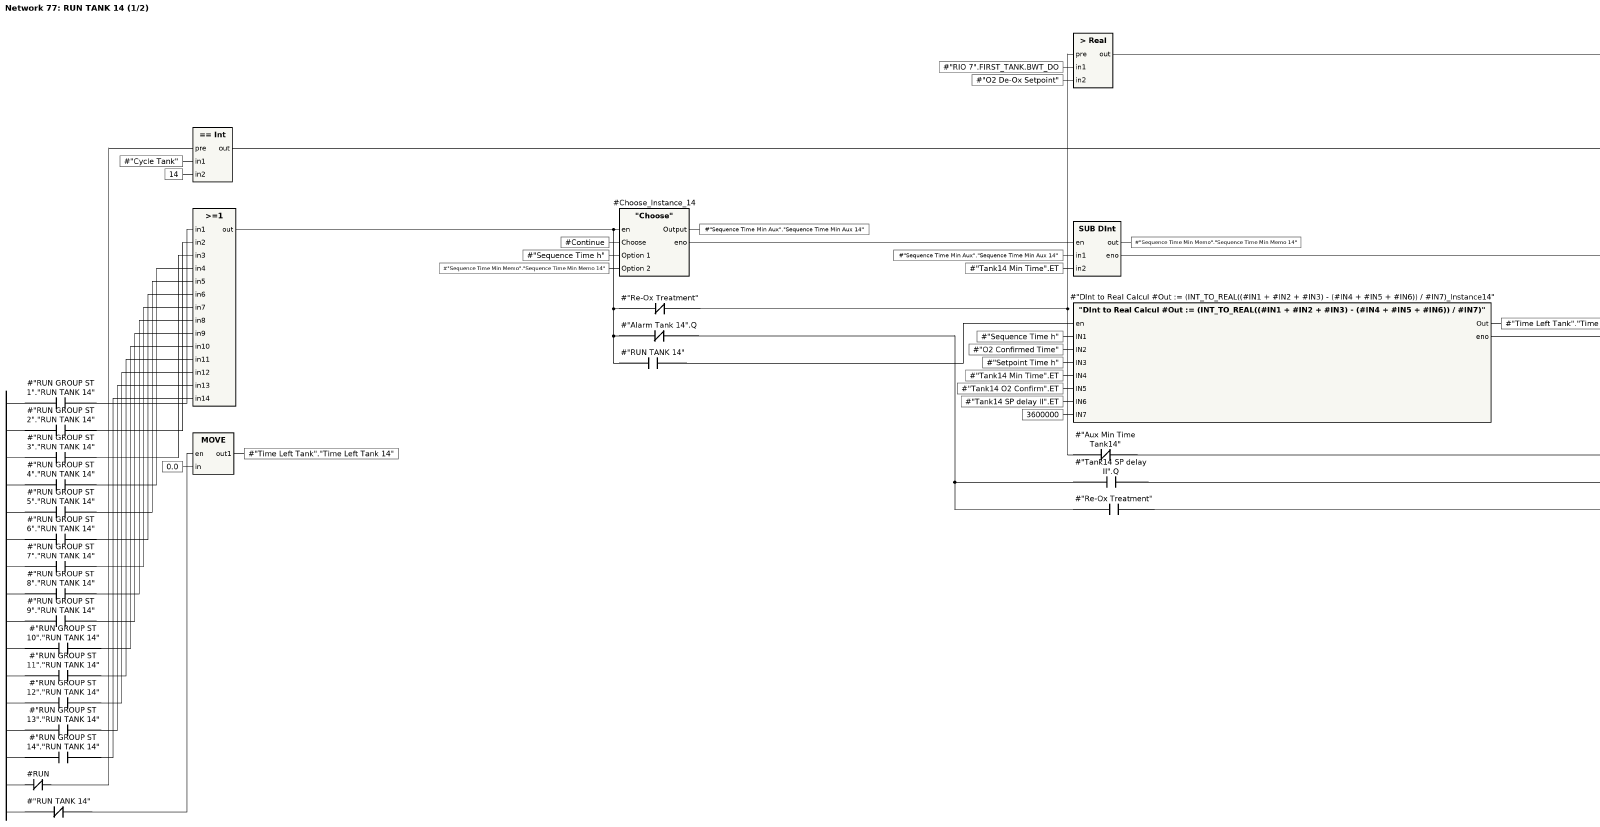
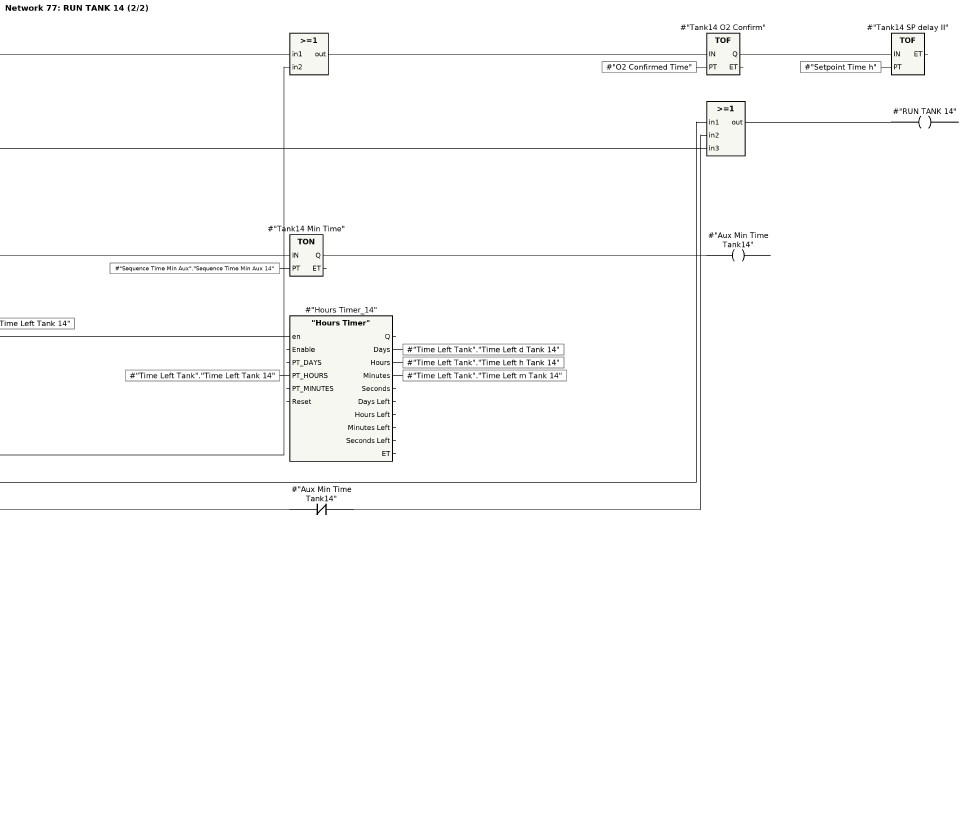
   #_w1 := #"RUN GROUP ST 1"."RUN TANK 14" OR #"RUN GROUP ST 2"."RUN TANK 14" OR #"RUN GROUP ST 3"."RUN TANK 14" OR #"RUN GROUP ST 4"."RUN TANK 14" OR #"RUN GROUP ST 5"."RUN TANK 14" OR #"RUN GROUP ST 6"."RUN TANK 14" OR #"RUN GROUP ST 7"."RUN TANK 14" OR #"RUN GROUP ST 8"."RUN TANK 14" OR #"RUN GROUP ST 9"."RUN TANK 14" OR #"RUN GROUP ST 10"."RUN TANK 14" OR #"RUN GROUP ST 11"."RUN TANK 14" OR #"RUN GROUP ST 12"."RUN TANK 14" OR #"RUN GROUP ST 13"."RUN TANK 14" OR #"RUN GROUP ST 14"."RUN TANK 14";
   #Choose_Instance_14(EN := #_w1,   // "Choose"
                       Choose := #Continue,
                       "Option 1" := #"Sequence Time h",
                       "Option 2" := #"Sequence Time Min Memo"."Sequence Time Min Memo 14",
                       Output => #"Sequence Time Min Aux"."Sequence Time Min Aux 14",
                       ENO => #_w2);
   IF #_w2 THEN
       #"Sequence Time Min Memo"."Sequence Time Min Memo 14" := #"Sequence Time Min Aux"."Sequence Time Min Aux 14" - #"Tank14 Min Time".ET;   // Memory of remained time for use to continue
   END_IF;
   #"Tank14 Min Time"(IN := #_w2, PT := #"Sequence Time Min Aux"."Sequence Time Min Aux 14");   // TON
   #"Aux Min Time Tank14" := #"Tank14 Min Time".Q;
   #"Tank14 O2 Confirm"(IN := #_w1 AND NOT #"Re-Ox Treatment" AND ((#"RIO 7".FIRST_TANK.BWT_DO > #"O2 De-Ox Setpoint") OR NOT #"Aux Min Time Tank14"),   // TOF
                        PT := #"O2 Confirmed Time");
   #"Tank14 SP delay II"(IN := #"Tank14 O2 Confirm".Q, PT := #"Setpoint Time h");   // TOF
   #"DInt to Real Calcul #Out := (INT_TO_REAL((#IN1 + #IN2 + #IN3) - (#IN4 + #IN5 + #IN6)) / #IN7)_Instance14"(EN := #_w1 AND #"RUN TANK 14",   // "DInt to Real Calcul #Out := (INT_TO_REAL((#IN1 + #IN2 + #IN3) - (#IN4 + #IN5 + #IN6)) / #IN7)"
                           IN1 := #"Sequence Time h",
                           IN2 := #"O2 Confirmed Time",
                           IN3 := #"Setpoint Time h",
                           IN4 := #"Tank14 Min Time".ET,
                           IN5 := #"Tank14 O2 Confirm".ET,
                           IN6 := #"Tank14 SP delay II".ET,
                           IN7 := 3600000,
                           Out => #"Time Left Tank"."Time Left Tank 14",
                           ENO => #_w3);
   IF #_w3 THEN
       #"Hours Timer_14"(PT_HOURS := #"Time Left Tank"."Time Left Tank 14",   // "Hours Timer"
                         Days => #"Time Left Tank"."Time Left d Tank 14",
                         Hours => #"Time Left Tank"."Time Left h Tank 14",
                         Minutes => #"Time Left Tank"."Time Left m Tank 14");
   END_IF;
   #"RUN TANK 14" := (#_w1 AND NOT #"Alarm Tank 14".Q AND (#"Tank14 SP delay II".Q OR (#"Re-Ox Treatment" AND NOT #"Aux Min Time Tank14"))) OR (NOT #RUN AND (#"Cycle Tank" = 14));
   IF NOT #"RUN TANK 14" THEN #"Time Left Tank"."Time Left Tank 14" := 0.0; END_IF;
END_REGION

REGION Network 78: RUN TANK 15
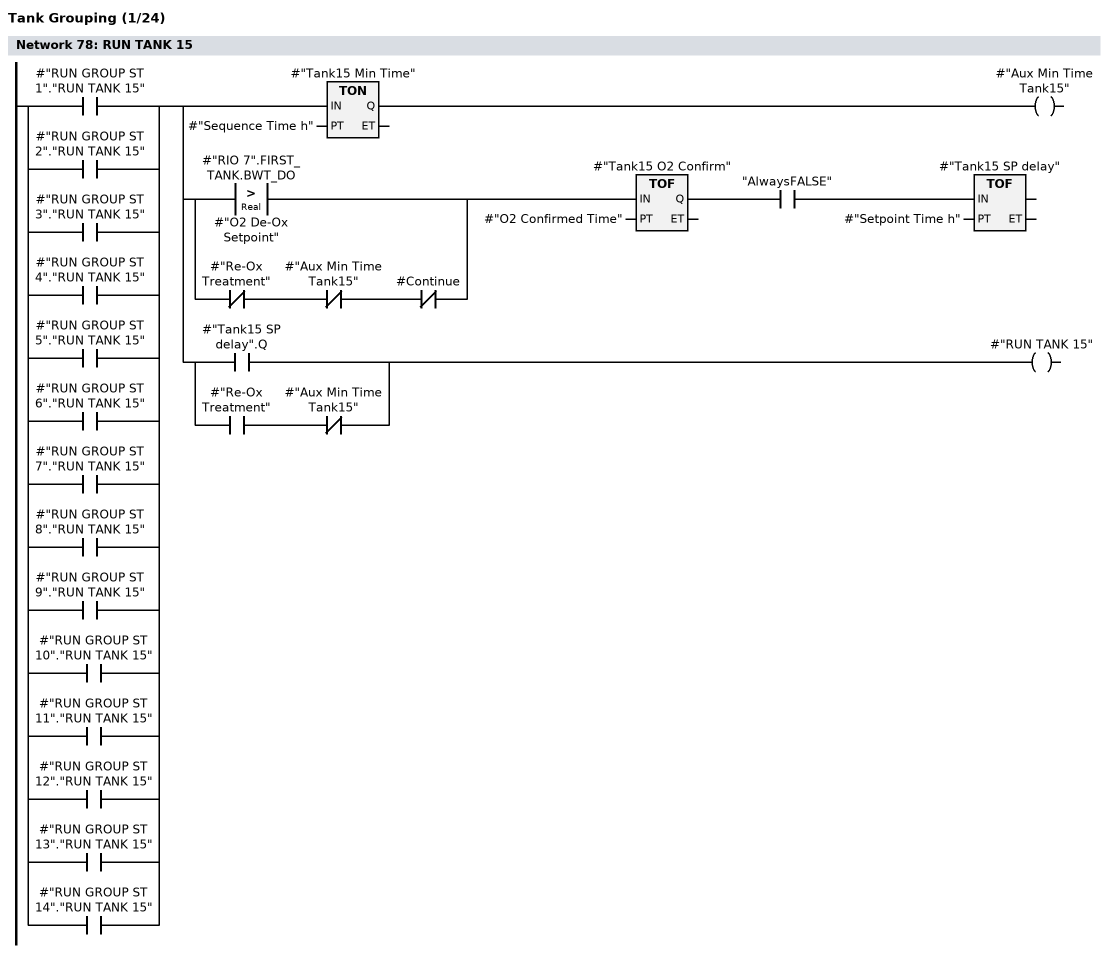
   #_w1 := #"RUN GROUP ST 1"."RUN TANK 15" OR #"RUN GROUP ST 2"."RUN TANK 15" OR #"RUN GROUP ST 3"."RUN TANK 15" OR #"RUN GROUP ST 4"."RUN TANK 15" OR #"RUN GROUP ST 5"."RUN TANK 15" OR #"RUN GROUP ST 6"."RUN TANK 15" OR #"RUN GROUP ST 7"."RUN TANK 15" OR #"RUN GROUP ST 8"."RUN TANK 15" OR #"RUN GROUP ST 9"."RUN TANK 15" OR #"RUN GROUP ST 10"."RUN TANK 15" OR #"RUN GROUP ST 11"."RUN TANK 15" OR #"RUN GROUP ST 12"."RUN TANK 15" OR #"RUN GROUP ST 13"."RUN TANK 15" OR #"RUN GROUP ST 14"."RUN TANK 15";
   #"Tank15 Min Time"(IN := #_w1, PT := #"Sequence Time h");   // TON
   #"Aux Min Time Tank15" := #"Tank15 Min Time".Q;
   #"Tank15 O2 Confirm"(IN := #_w1 AND ((#"RIO 7".FIRST_TANK.BWT_DO > #"O2 De-Ox Setpoint") OR (NOT #"Re-Ox Treatment" AND NOT #"Aux Min Time Tank15" AND NOT #Continue)),   // TOF
                        PT := #"O2 Confirmed Time");
   #"Tank15 SP delay"(IN := #"Tank15 O2 Confirm".Q AND "AlwaysFALSE", PT := #"Setpoint Time h");   // TOF
   #"RUN TANK 15" := #_w1 AND (#"Tank15 SP delay".Q OR (#"Re-Ox Treatment" AND NOT #"Aux Min Time Tank15"));
END_REGION

REGION Network 79: RUN TANK 16
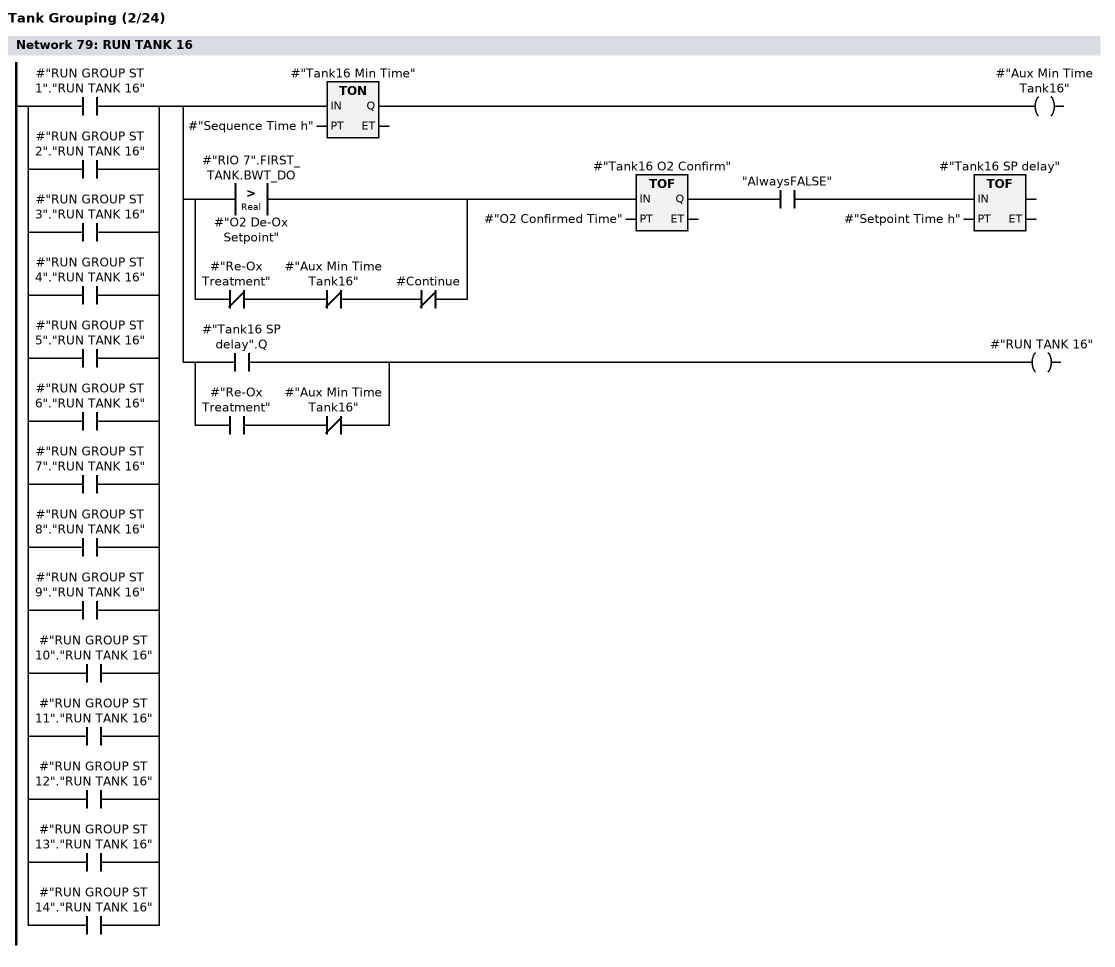
   #_w1 := #"RUN GROUP ST 1"."RUN TANK 16" OR #"RUN GROUP ST 2"."RUN TANK 16" OR #"RUN GROUP ST 3"."RUN TANK 16" OR #"RUN GROUP ST 4"."RUN TANK 16" OR #"RUN GROUP ST 5"."RUN TANK 16" OR #"RUN GROUP ST 6"."RUN TANK 16" OR #"RUN GROUP ST 7"."RUN TANK 16" OR #"RUN GROUP ST 8"."RUN TANK 16" OR #"RUN GROUP ST 9"."RUN TANK 16" OR #"RUN GROUP ST 10"."RUN TANK 16" OR #"RUN GROUP ST 11"."RUN TANK 16" OR #"RUN GROUP ST 12"."RUN TANK 16" OR #"RUN GROUP ST 13"."RUN TANK 16" OR #"RUN GROUP ST 14"."RUN TANK 16";
   #"Tank16 Min Time"(IN := #_w1, PT := #"Sequence Time h");   // TON
   #"Aux Min Time Tank16" := #"Tank16 Min Time".Q;
   #"Tank16 O2 Confirm"(IN := #_w1 AND ((#"RIO 7".FIRST_TANK.BWT_DO > #"O2 De-Ox Setpoint") OR (NOT #"Re-Ox Treatment" AND NOT #"Aux Min Time Tank16" AND NOT #Continue)),   // TOF
                        PT := #"O2 Confirmed Time");
   #"Tank16 SP delay"(IN := #"Tank16 O2 Confirm".Q AND "AlwaysFALSE", PT := #"Setpoint Time h");   // TOF
   #"RUN TANK 16" := #_w1 AND (#"Tank16 SP delay".Q OR (#"Re-Ox Treatment" AND NOT #"Aux Min Time Tank16"));
END_REGION

REGION Network 80: RUN TANK 17
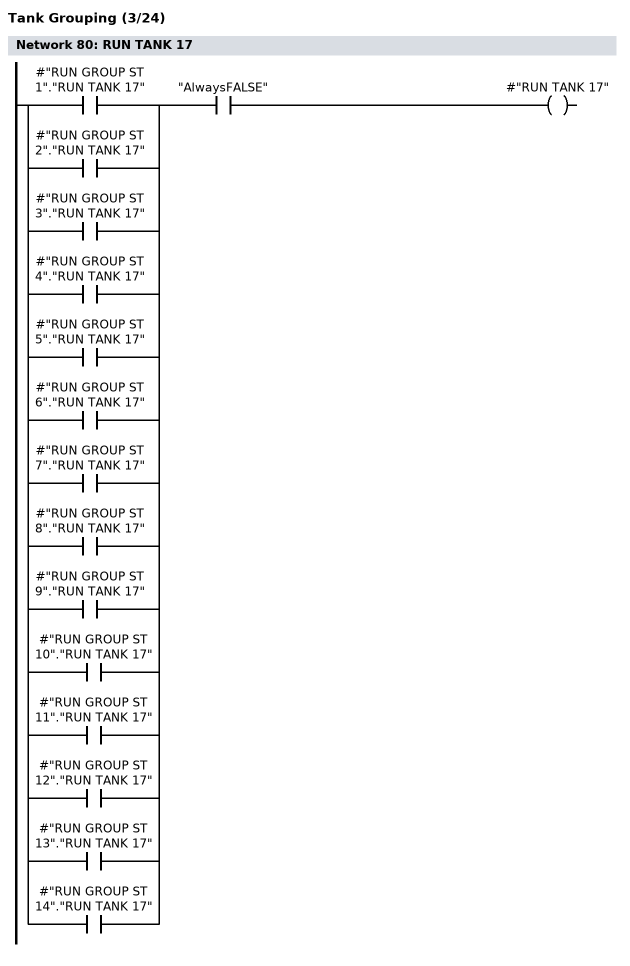
   RUNG wire#powerrail
      Contact( #"RUN GROUP ST 1"."RUN TANK 17" )
      wire#w1
      Contact( "AlwaysFALSE" )
      Coil( #"RUN TANK 17" )
   END_RUNG
   RUNG wire#powerrail
      Contact( #"RUN GROUP ST 2"."RUN TANK 17" )
   END_RUNG wire#w1
   RUNG wire#powerrail
      Contact( #"RUN GROUP ST 3"."RUN TANK 17" )
   END_RUNG wire#w1
   RUNG wire#powerrail
      Contact( #"RUN GROUP ST 4"."RUN TANK 17" )
   END_RUNG wire#w1
   RUNG wire#powerrail
      Contact( #"RUN GROUP ST 5"."RUN TANK 17" )
   END_RUNG wire#w1
   RUNG wire#powerrail
      Contact( #"RUN GROUP ST 6"."RUN TANK 17" )
   END_RUNG wire#w1
   RUNG wire#powerrail
      Contact( #"RUN GROUP ST 7"."RUN TANK 17" )
   END_RUNG wire#w1
   RUNG wire#powerrail
      Contact( #"RUN GROUP ST 8"."RUN TANK 17" )
   END_RUNG wire#w1
   RUNG wire#powerrail
      Contact( #"RUN GROUP ST 9"."RUN TANK 17" )
   END_RUNG wire#w1
   RUNG wire#powerrail
      Contact( #"RUN GROUP ST 10"."RUN TANK 17" )
   END_RUNG wire#w1
   RUNG wire#powerrail
      Contact( #"RUN GROUP ST 11"."RUN TANK 17" )
   END_RUNG wire#w1
   RUNG wire#powerrail
      Contact( #"RUN GROUP ST 12"."RUN TANK 17" )
   END_RUNG wire#w1
   RUNG wire#powerrail
      Contact( #"RUN GROUP ST 13"."RUN TANK 17" )
   END_RUNG wire#w1
   RUNG wire#powerrail
      Contact( #"RUN GROUP ST 14"."RUN TANK 17" )
   END_RUNG wire#w1
   // the same network as SCL:
   #"RUN TANK 17" := (#"RUN GROUP ST 1"."RUN TANK 17" OR #"RUN GROUP ST 2"."RUN TANK 17" OR #"RUN GROUP ST 3"."RUN TANK 17" OR #"RUN GROUP ST 4"."RUN TANK 17" OR #"RUN GROUP ST 5"."RUN TANK 17" OR #"RUN GROUP ST 6"."RUN TANK 17" OR #"RUN GROUP ST 7"."RUN TANK 17" OR #"RUN GROUP ST 8"."RUN TANK 17" OR #"RUN GROUP ST 9"."RUN TANK 17" OR #"RUN GROUP ST 10"."RUN TANK 17" OR #"RUN GROUP ST 11"."RUN TANK 17" OR #"RUN GROUP ST 12"."RUN TANK 17" OR #"RUN GROUP ST 13"."RUN TANK 17" OR #"RUN GROUP ST 14"."RUN TANK 17") AND "AlwaysFALSE";
END_REGION

REGION Network 81: RUN TANK 18
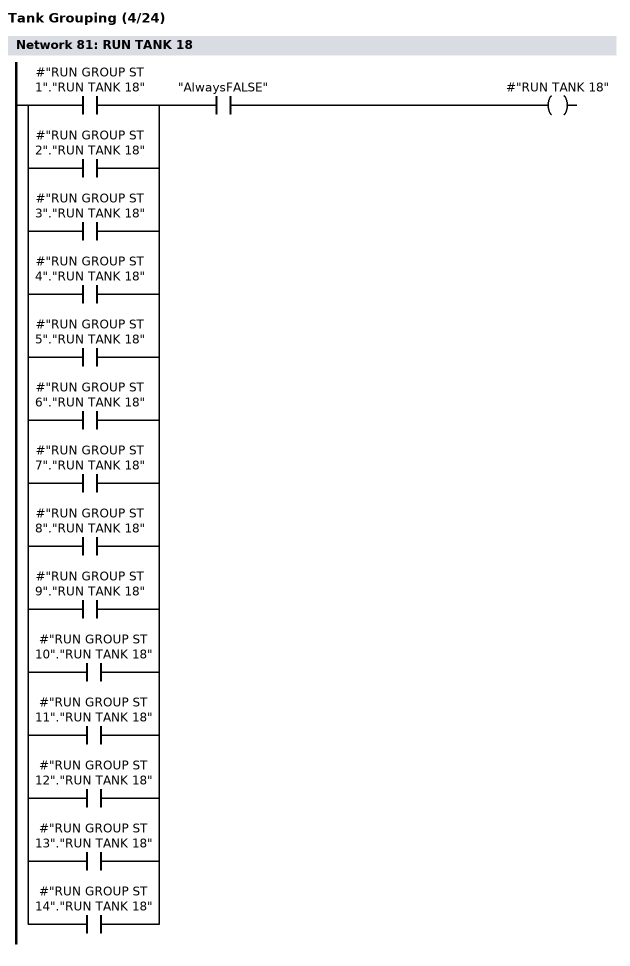
   RUNG wire#powerrail
      Contact( #"RUN GROUP ST 1"."RUN TANK 18" )
      wire#w1
      Contact( "AlwaysFALSE" )
      Coil( #"RUN TANK 18" )
   END_RUNG
   RUNG wire#powerrail
      Contact( #"RUN GROUP ST 2"."RUN TANK 18" )
   END_RUNG wire#w1
   RUNG wire#powerrail
      Contact( #"RUN GROUP ST 3"."RUN TANK 18" )
   END_RUNG wire#w1
   RUNG wire#powerrail
      Contact( #"RUN GROUP ST 4"."RUN TANK 18" )
   END_RUNG wire#w1
   RUNG wire#powerrail
      Contact( #"RUN GROUP ST 5"."RUN TANK 18" )
   END_RUNG wire#w1
   RUNG wire#powerrail
      Contact( #"RUN GROUP ST 6"."RUN TANK 18" )
   END_RUNG wire#w1
   RUNG wire#powerrail
      Contact( #"RUN GROUP ST 7"."RUN TANK 18" )
   END_RUNG wire#w1
   RUNG wire#powerrail
      Contact( #"RUN GROUP ST 8"."RUN TANK 18" )
   END_RUNG wire#w1
   RUNG wire#powerrail
      Contact( #"RUN GROUP ST 9"."RUN TANK 18" )
   END_RUNG wire#w1
   RUNG wire#powerrail
      Contact( #"RUN GROUP ST 10"."RUN TANK 18" )
   END_RUNG wire#w1
   RUNG wire#powerrail
      Contact( #"RUN GROUP ST 11"."RUN TANK 18" )
   END_RUNG wire#w1
   RUNG wire#powerrail
      Contact( #"RUN GROUP ST 12"."RUN TANK 18" )
   END_RUNG wire#w1
   RUNG wire#powerrail
      Contact( #"RUN GROUP ST 13"."RUN TANK 18" )
   END_RUNG wire#w1
   RUNG wire#powerrail
      Contact( #"RUN GROUP ST 14"."RUN TANK 18" )
   END_RUNG wire#w1
   // the same network as SCL:
   #"RUN TANK 18" := (#"RUN GROUP ST 1"."RUN TANK 18" OR #"RUN GROUP ST 2"."RUN TANK 18" OR #"RUN GROUP ST 3"."RUN TANK 18" OR #"RUN GROUP ST 4"."RUN TANK 18" OR #"RUN GROUP ST 5"."RUN TANK 18" OR #"RUN GROUP ST 6"."RUN TANK 18" OR #"RUN GROUP ST 7"."RUN TANK 18" OR #"RUN GROUP ST 8"."RUN TANK 18" OR #"RUN GROUP ST 9"."RUN TANK 18" OR #"RUN GROUP ST 10"."RUN TANK 18" OR #"RUN GROUP ST 11"."RUN TANK 18" OR #"RUN GROUP ST 12"."RUN TANK 18" OR #"RUN GROUP ST 13"."RUN TANK 18" OR #"RUN GROUP ST 14"."RUN TANK 18") AND "AlwaysFALSE";
END_REGION

REGION Network 82: RUN TANK 19
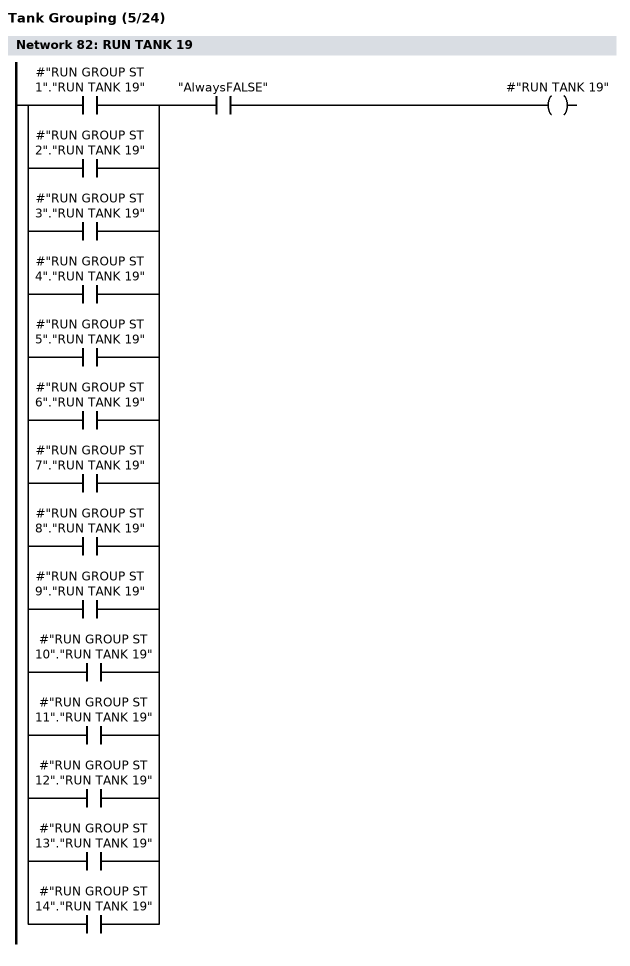
   RUNG wire#powerrail
      Contact( #"RUN GROUP ST 1"."RUN TANK 19" )
      wire#w1
      Contact( "AlwaysFALSE" )
      Coil( #"RUN TANK 19" )
   END_RUNG
   RUNG wire#powerrail
      Contact( #"RUN GROUP ST 2"."RUN TANK 19" )
   END_RUNG wire#w1
   RUNG wire#powerrail
      Contact( #"RUN GROUP ST 3"."RUN TANK 19" )
   END_RUNG wire#w1
   RUNG wire#powerrail
      Contact( #"RUN GROUP ST 4"."RUN TANK 19" )
   END_RUNG wire#w1
   RUNG wire#powerrail
      Contact( #"RUN GROUP ST 5"."RUN TANK 19" )
   END_RUNG wire#w1
   RUNG wire#powerrail
      Contact( #"RUN GROUP ST 6"."RUN TANK 19" )
   END_RUNG wire#w1
   RUNG wire#powerrail
      Contact( #"RUN GROUP ST 7"."RUN TANK 19" )
   END_RUNG wire#w1
   RUNG wire#powerrail
      Contact( #"RUN GROUP ST 8"."RUN TANK 19" )
   END_RUNG wire#w1
   RUNG wire#powerrail
      Contact( #"RUN GROUP ST 9"."RUN TANK 19" )
   END_RUNG wire#w1
   RUNG wire#powerrail
      Contact( #"RUN GROUP ST 10"."RUN TANK 19" )
   END_RUNG wire#w1
   RUNG wire#powerrail
      Contact( #"RUN GROUP ST 11"."RUN TANK 19" )
   END_RUNG wire#w1
   RUNG wire#powerrail
      Contact( #"RUN GROUP ST 12"."RUN TANK 19" )
   END_RUNG wire#w1
   RUNG wire#powerrail
      Contact( #"RUN GROUP ST 13"."RUN TANK 19" )
   END_RUNG wire#w1
   RUNG wire#powerrail
      Contact( #"RUN GROUP ST 14"."RUN TANK 19" )
   END_RUNG wire#w1
   // the same network as SCL:
   #"RUN TANK 19" := (#"RUN GROUP ST 1"."RUN TANK 19" OR #"RUN GROUP ST 2"."RUN TANK 19" OR #"RUN GROUP ST 3"."RUN TANK 19" OR #"RUN GROUP ST 4"."RUN TANK 19" OR #"RUN GROUP ST 5"."RUN TANK 19" OR #"RUN GROUP ST 6"."RUN TANK 19" OR #"RUN GROUP ST 7"."RUN TANK 19" OR #"RUN GROUP ST 8"."RUN TANK 19" OR #"RUN GROUP ST 9"."RUN TANK 19" OR #"RUN GROUP ST 10"."RUN TANK 19" OR #"RUN GROUP ST 11"."RUN TANK 19" OR #"RUN GROUP ST 12"."RUN TANK 19" OR #"RUN GROUP ST 13"."RUN TANK 19" OR #"RUN GROUP ST 14"."RUN TANK 19") AND "AlwaysFALSE";
END_REGION

REGION Network 83: RUN TANK 20
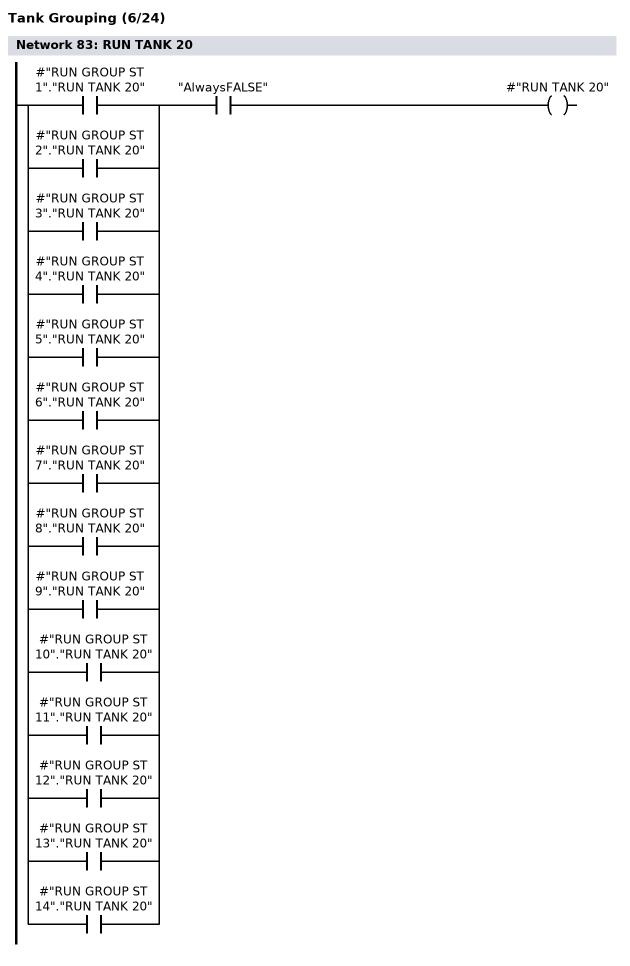
   RUNG wire#powerrail
      Contact( #"RUN GROUP ST 1"."RUN TANK 20" )
      wire#w1
      Contact( "AlwaysFALSE" )
      Coil( #"RUN TANK 20" )
   END_RUNG
   RUNG wire#powerrail
      Contact( #"RUN GROUP ST 2"."RUN TANK 20" )
   END_RUNG wire#w1
   RUNG wire#powerrail
      Contact( #"RUN GROUP ST 3"."RUN TANK 20" )
   END_RUNG wire#w1
   RUNG wire#powerrail
      Contact( #"RUN GROUP ST 4"."RUN TANK 20" )
   END_RUNG wire#w1
   RUNG wire#powerrail
      Contact( #"RUN GROUP ST 5"."RUN TANK 20" )
   END_RUNG wire#w1
   RUNG wire#powerrail
      Contact( #"RUN GROUP ST 6"."RUN TANK 20" )
   END_RUNG wire#w1
   RUNG wire#powerrail
      Contact( #"RUN GROUP ST 7"."RUN TANK 20" )
   END_RUNG wire#w1
   RUNG wire#powerrail
      Contact( #"RUN GROUP ST 8"."RUN TANK 20" )
   END_RUNG wire#w1
   RUNG wire#powerrail
      Contact( #"RUN GROUP ST 9"."RUN TANK 20" )
   END_RUNG wire#w1
   RUNG wire#powerrail
      Contact( #"RUN GROUP ST 10"."RUN TANK 20" )
   END_RUNG wire#w1
   RUNG wire#powerrail
      Contact( #"RUN GROUP ST 11"."RUN TANK 20" )
   END_RUNG wire#w1
   RUNG wire#powerrail
      Contact( #"RUN GROUP ST 12"."RUN TANK 20" )
   END_RUNG wire#w1
   RUNG wire#powerrail
      Contact( #"RUN GROUP ST 13"."RUN TANK 20" )
   END_RUNG wire#w1
   RUNG wire#powerrail
      Contact( #"RUN GROUP ST 14"."RUN TANK 20" )
   END_RUNG wire#w1
   // the same network as SCL:
   #"RUN TANK 20" := (#"RUN GROUP ST 1"."RUN TANK 20" OR #"RUN GROUP ST 2"."RUN TANK 20" OR #"RUN GROUP ST 3"."RUN TANK 20" OR #"RUN GROUP ST 4"."RUN TANK 20" OR #"RUN GROUP ST 5"."RUN TANK 20" OR #"RUN GROUP ST 6"."RUN TANK 20" OR #"RUN GROUP ST 7"."RUN TANK 20" OR #"RUN GROUP ST 8"."RUN TANK 20" OR #"RUN GROUP ST 9"."RUN TANK 20" OR #"RUN GROUP ST 10"."RUN TANK 20" OR #"RUN GROUP ST 11"."RUN TANK 20" OR #"RUN GROUP ST 12"."RUN TANK 20" OR #"RUN GROUP ST 13"."RUN TANK 20" OR #"RUN GROUP ST 14"."RUN TANK 20") AND "AlwaysFALSE";
END_REGION

REGION Network 84: RUN TANK 21
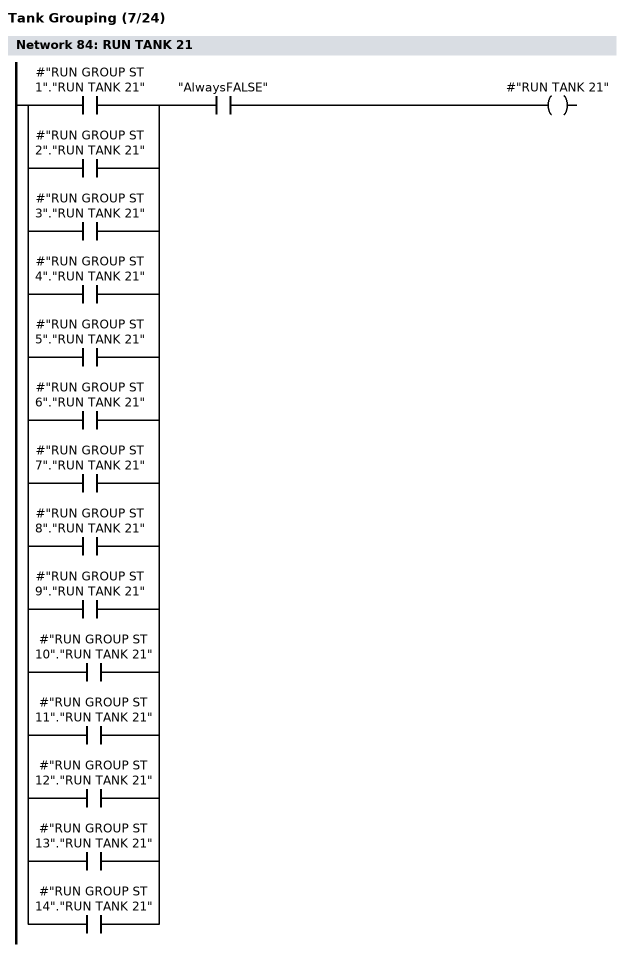
   RUNG wire#powerrail
      Contact( #"RUN GROUP ST 1"."RUN TANK 21" )
      wire#w1
      Contact( "AlwaysFALSE" )
      Coil( #"RUN TANK 21" )
   END_RUNG
   RUNG wire#powerrail
      Contact( #"RUN GROUP ST 2"."RUN TANK 21" )
   END_RUNG wire#w1
   RUNG wire#powerrail
      Contact( #"RUN GROUP ST 3"."RUN TANK 21" )
   END_RUNG wire#w1
   RUNG wire#powerrail
      Contact( #"RUN GROUP ST 4"."RUN TANK 21" )
   END_RUNG wire#w1
   RUNG wire#powerrail
      Contact( #"RUN GROUP ST 5"."RUN TANK 21" )
   END_RUNG wire#w1
   RUNG wire#powerrail
      Contact( #"RUN GROUP ST 6"."RUN TANK 21" )
   END_RUNG wire#w1
   RUNG wire#powerrail
      Contact( #"RUN GROUP ST 7"."RUN TANK 21" )
   END_RUNG wire#w1
   RUNG wire#powerrail
      Contact( #"RUN GROUP ST 8"."RUN TANK 21" )
   END_RUNG wire#w1
   RUNG wire#powerrail
      Contact( #"RUN GROUP ST 9"."RUN TANK 21" )
   END_RUNG wire#w1
   RUNG wire#powerrail
      Contact( #"RUN GROUP ST 10"."RUN TANK 21" )
   END_RUNG wire#w1
   RUNG wire#powerrail
      Contact( #"RUN GROUP ST 11"."RUN TANK 21" )
   END_RUNG wire#w1
   RUNG wire#powerrail
      Contact( #"RUN GROUP ST 12"."RUN TANK 21" )
   END_RUNG wire#w1
   RUNG wire#powerrail
      Contact( #"RUN GROUP ST 13"."RUN TANK 21" )
   END_RUNG wire#w1
   RUNG wire#powerrail
      Contact( #"RUN GROUP ST 14"."RUN TANK 21" )
   END_RUNG wire#w1
   // the same network as SCL:
   #"RUN TANK 21" := (#"RUN GROUP ST 1"."RUN TANK 21" OR #"RUN GROUP ST 2"."RUN TANK 21" OR #"RUN GROUP ST 3"."RUN TANK 21" OR #"RUN GROUP ST 4"."RUN TANK 21" OR #"RUN GROUP ST 5"."RUN TANK 21" OR #"RUN GROUP ST 6"."RUN TANK 21" OR #"RUN GROUP ST 7"."RUN TANK 21" OR #"RUN GROUP ST 8"."RUN TANK 21" OR #"RUN GROUP ST 9"."RUN TANK 21" OR #"RUN GROUP ST 10"."RUN TANK 21" OR #"RUN GROUP ST 11"."RUN TANK 21" OR #"RUN GROUP ST 12"."RUN TANK 21" OR #"RUN GROUP ST 13"."RUN TANK 21" OR #"RUN GROUP ST 14"."RUN TANK 21") AND "AlwaysFALSE";
END_REGION

REGION Network 85: RUN TANK 22
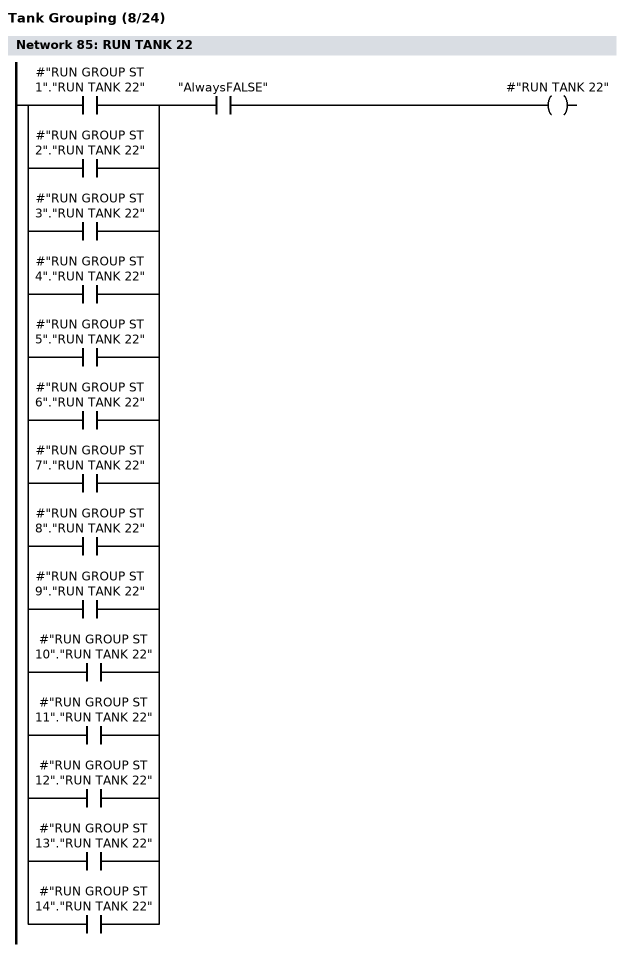
   RUNG wire#powerrail
      Contact( #"RUN GROUP ST 1"."RUN TANK 22" )
      wire#w1
      Contact( "AlwaysFALSE" )
      Coil( #"RUN TANK 22" )
   END_RUNG
   RUNG wire#powerrail
      Contact( #"RUN GROUP ST 2"."RUN TANK 22" )
   END_RUNG wire#w1
   RUNG wire#powerrail
      Contact( #"RUN GROUP ST 3"."RUN TANK 22" )
   END_RUNG wire#w1
   RUNG wire#powerrail
      Contact( #"RUN GROUP ST 4"."RUN TANK 22" )
   END_RUNG wire#w1
   RUNG wire#powerrail
      Contact( #"RUN GROUP ST 5"."RUN TANK 22" )
   END_RUNG wire#w1
   RUNG wire#powerrail
      Contact( #"RUN GROUP ST 6"."RUN TANK 22" )
   END_RUNG wire#w1
   RUNG wire#powerrail
      Contact( #"RUN GROUP ST 7"."RUN TANK 22" )
   END_RUNG wire#w1
   RUNG wire#powerrail
      Contact( #"RUN GROUP ST 8"."RUN TANK 22" )
   END_RUNG wire#w1
   RUNG wire#powerrail
      Contact( #"RUN GROUP ST 9"."RUN TANK 22" )
   END_RUNG wire#w1
   RUNG wire#powerrail
      Contact( #"RUN GROUP ST 10"."RUN TANK 22" )
   END_RUNG wire#w1
   RUNG wire#powerrail
      Contact( #"RUN GROUP ST 11"."RUN TANK 22" )
   END_RUNG wire#w1
   RUNG wire#powerrail
      Contact( #"RUN GROUP ST 12"."RUN TANK 22" )
   END_RUNG wire#w1
   RUNG wire#powerrail
      Contact( #"RUN GROUP ST 13"."RUN TANK 22" )
   END_RUNG wire#w1
   RUNG wire#powerrail
      Contact( #"RUN GROUP ST 14"."RUN TANK 22" )
   END_RUNG wire#w1
   // the same network as SCL:
   #"RUN TANK 22" := (#"RUN GROUP ST 1"."RUN TANK 22" OR #"RUN GROUP ST 2"."RUN TANK 22" OR #"RUN GROUP ST 3"."RUN TANK 22" OR #"RUN GROUP ST 4"."RUN TANK 22" OR #"RUN GROUP ST 5"."RUN TANK 22" OR #"RUN GROUP ST 6"."RUN TANK 22" OR #"RUN GROUP ST 7"."RUN TANK 22" OR #"RUN GROUP ST 8"."RUN TANK 22" OR #"RUN GROUP ST 9"."RUN TANK 22" OR #"RUN GROUP ST 10"."RUN TANK 22" OR #"RUN GROUP ST 11"."RUN TANK 22" OR #"RUN GROUP ST 12"."RUN TANK 22" OR #"RUN GROUP ST 13"."RUN TANK 22" OR #"RUN GROUP ST 14"."RUN TANK 22") AND "AlwaysFALSE";
END_REGION

REGION Network 86: RUN TANK 23
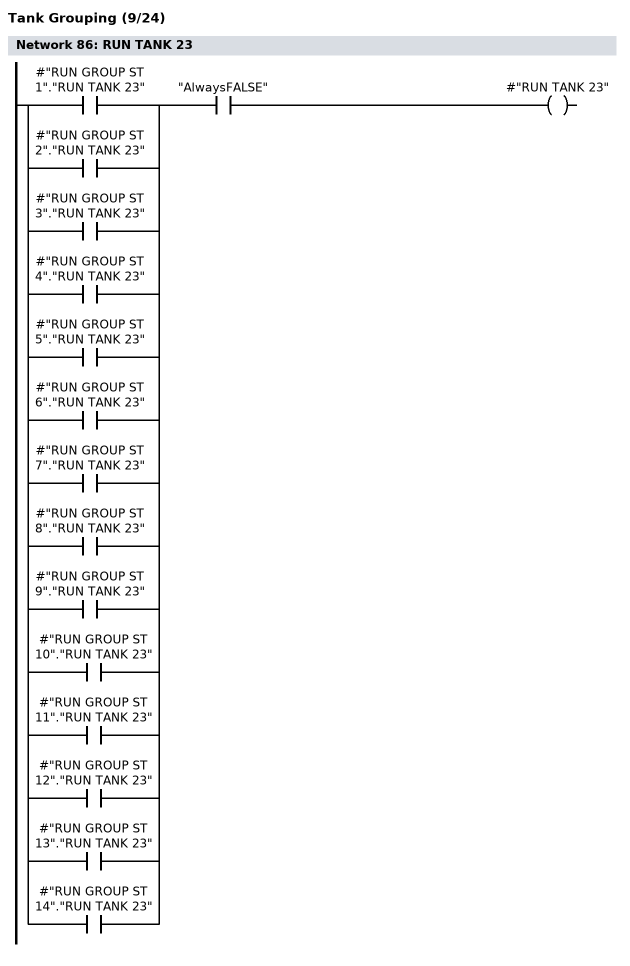
   RUNG wire#powerrail
      Contact( #"RUN GROUP ST 1"."RUN TANK 23" )
      wire#w1
      Contact( "AlwaysFALSE" )
      Coil( #"RUN TANK 23" )
   END_RUNG
   RUNG wire#powerrail
      Contact( #"RUN GROUP ST 2"."RUN TANK 23" )
   END_RUNG wire#w1
   RUNG wire#powerrail
      Contact( #"RUN GROUP ST 3"."RUN TANK 23" )
   END_RUNG wire#w1
   RUNG wire#powerrail
      Contact( #"RUN GROUP ST 4"."RUN TANK 23" )
   END_RUNG wire#w1
   RUNG wire#powerrail
      Contact( #"RUN GROUP ST 5"."RUN TANK 23" )
   END_RUNG wire#w1
   RUNG wire#powerrail
      Contact( #"RUN GROUP ST 6"."RUN TANK 23" )
   END_RUNG wire#w1
   RUNG wire#powerrail
      Contact( #"RUN GROUP ST 7"."RUN TANK 23" )
   END_RUNG wire#w1
   RUNG wire#powerrail
      Contact( #"RUN GROUP ST 8"."RUN TANK 23" )
   END_RUNG wire#w1
   RUNG wire#powerrail
      Contact( #"RUN GROUP ST 9"."RUN TANK 23" )
   END_RUNG wire#w1
   RUNG wire#powerrail
      Contact( #"RUN GROUP ST 10"."RUN TANK 23" )
   END_RUNG wire#w1
   RUNG wire#powerrail
      Contact( #"RUN GROUP ST 11"."RUN TANK 23" )
   END_RUNG wire#w1
   RUNG wire#powerrail
      Contact( #"RUN GROUP ST 12"."RUN TANK 23" )
   END_RUNG wire#w1
   RUNG wire#powerrail
      Contact( #"RUN GROUP ST 13"."RUN TANK 23" )
   END_RUNG wire#w1
   RUNG wire#powerrail
      Contact( #"RUN GROUP ST 14"."RUN TANK 23" )
   END_RUNG wire#w1
   // the same network as SCL:
   #"RUN TANK 23" := (#"RUN GROUP ST 1"."RUN TANK 23" OR #"RUN GROUP ST 2"."RUN TANK 23" OR #"RUN GROUP ST 3"."RUN TANK 23" OR #"RUN GROUP ST 4"."RUN TANK 23" OR #"RUN GROUP ST 5"."RUN TANK 23" OR #"RUN GROUP ST 6"."RUN TANK 23" OR #"RUN GROUP ST 7"."RUN TANK 23" OR #"RUN GROUP ST 8"."RUN TANK 23" OR #"RUN GROUP ST 9"."RUN TANK 23" OR #"RUN GROUP ST 10"."RUN TANK 23" OR #"RUN GROUP ST 11"."RUN TANK 23" OR #"RUN GROUP ST 12"."RUN TANK 23" OR #"RUN GROUP ST 13"."RUN TANK 23" OR #"RUN GROUP ST 14"."RUN TANK 23") AND "AlwaysFALSE";
END_REGION

REGION Network 87: RUN TANK 24